// TIA Portal project "EEEB EMBU 4_V17" (V17) (continued)
VERSION : 0.1
   VAR
      "CONNECT-MGE-PCM-E-CF-01" : TCON_IP_v4;   // Dados de configuração
      "CONNECT-MGE-QGBT-AUX-01" : TCON_IP_v4;   // Dados de configuração
      "Register-MGE-PCM-E-CF-01" : Array[0..38] of DInt;   // Tabela para receber os dados
      "Register-MGE-QGBT-AUX-01" : Array[0..38] of DInt;   // Tabela para receber os dados
      LADDR_PROFINET : Hw_IoSystem := 261;   // Endereço de hardware
      MODE_PROFINET : UInt := 4;   // Modo de operação da funcção
      RET_VAL_PROFINET : Int;   // Terorno de diagnóstico
      ESTADO_PROFINET : Array[0..1023] of Bool;   // Diagnóstico da rede PROFINET
      DONE_MB : Array[0..60] of Bool;   // Sinaliza fim de execução
      BUSY_MB : Array[0..60] of Bool;   // Sinaliza espera
      ERROR_MB : Array[0..60] of Bool;   // Sinaliza erro
      STATUS_MB : Array[0..60] of Word;   // Satus da comunicação
      START_MB : Array[0..60] of Bool;   // Inicia comunicação
      FCOM_MB : Array[0..60] of Bool;   // Falha de comunicação
      HAB_MB : Array[0..60] of Bool;   // Habilita comunicação MODBUS
      INICIA_MB : Bool;   // INICIA CICLO DE COMUNICAÇÃO MODBUS
      INI_AUX_MB : Bool;   // AUXILIAR DE INICIALIZAÇÃO
   END_VAR
BEGIN
   "CONNECT-MGE-PCM-E-CF-01".LocalPort := 0;
   "CONNECT-MGE-PCM-E-CF-01".RemotePort := 502;
   "CONNECT-MGE-PCM-E-CF-01".RemoteAddress.ADDR[4] := 59;
   "CONNECT-MGE-PCM-E-CF-01".RemoteAddress.ADDR[3] := 2;
   "CONNECT-MGE-PCM-E-CF-01".RemoteAddress.ADDR[2] := 168;
   "CONNECT-MGE-PCM-E-CF-01".RemoteAddress.ADDR[1] := 192;
   "CONNECT-MGE-PCM-E-CF-01".ActiveEstablished := TRUE;
   "CONNECT-MGE-PCM-E-CF-01".ConnectionType := 11;
   "CONNECT-MGE-PCM-E-CF-01".ID := 10;
   "CONNECT-MGE-PCM-E-CF-01".InterfaceId := 64;
   "CONNECT-MGE-QGBT-AUX-01".LocalPort := 0;
   "CONNECT-MGE-QGBT-AUX-01".RemotePort := 502;
   "CONNECT-MGE-QGBT-AUX-01".RemoteAddress.ADDR[4] := 59;
   "CONNECT-MGE-QGBT-AUX-01".RemoteAddress.ADDR[3] := 2;
   "CONNECT-MGE-QGBT-AUX-01".RemoteAddress.ADDR[2] := 168;
   "CONNECT-MGE-QGBT-AUX-01".RemoteAddress.ADDR[1] := 192;
   "CONNECT-MGE-QGBT-AUX-01".ActiveEstablished := TRUE;
   "CONNECT-MGE-QGBT-AUX-01".ConnectionType := 11;
   "CONNECT-MGE-QGBT-AUX-01".ID := 10;
   "CONNECT-MGE-QGBT-AUX-01".InterfaceId := 64;
   // "Register-MGE-PCM-E-CF-01"[0] : Tensão (L-N) fase 1
   // "Register-MGE-PCM-E-CF-01"[1] : Tensão (L-L) fase 1-2
   // "Register-MGE-PCM-E-CF-01"[2] : Corrente fase 1
   // "Register-MGE-PCM-E-CF-01"[3] : Cos φ fase 1
   // "Register-MGE-PCM-E-CF-01"[4] : Fator de potencia fase 1
   // "Register-MGE-PCM-E-CF-01"[5] : Potencia ativa fase 1
   // "Register-MGE-PCM-E-CF-01"[6] : Potência reativa fase 1
   // "Register-MGE-PCM-E-CF-01"[7] : Potência aparente fase 1
   // "Register-MGE-PCM-E-CF-01"[8] : THDV fase 1
   // "Register-MGE-PCM-E-CF-01"[9] : THDI fase 1
   // "Register-MGE-PCM-E-CF-01"[10] : Tensão (L-N) fase 2
   // "Register-MGE-PCM-E-CF-01"[11] : Tensão (L-L) fase 2-3
   // "Register-MGE-PCM-E-CF-01"[12] : Corrente fase 2
   // "Register-MGE-PCM-E-CF-01"[13] : Cos φ fase 2
   // "Register-MGE-PCM-E-CF-01"[14] : Fator de potência fase 2
   // "Register-MGE-PCM-E-CF-01"[15] : Potência ativa fase 2
   // "Register-MGE-PCM-E-CF-01"[16] : Potência reativa fase 2
   // "Register-MGE-PCM-E-CF-01"[17] : Potência aparente fase 2
   // "Register-MGE-PCM-E-CF-01"[18] : THDV fase 2
   // "Register-MGE-PCM-E-CF-01"[19] : THDI fase 2
   // "Register-MGE-PCM-E-CF-01"[20] : Tensão (L-N) fase 3
   // "Register-MGE-PCM-E-CF-01"[21] : Tensão (L-L) fase 3-1
   // "Register-MGE-PCM-E-CF-01"[22] : Corrente fase 3
   // "Register-MGE-PCM-E-CF-01"[23] : Cos φ fase 3
   // "Register-MGE-PCM-E-CF-01"[24] : Fator de potência fase 3
   // "Register-MGE-PCM-E-CF-01"[25] : Potência ativa fase 3
   // "Register-MGE-PCM-E-CF-01"[26] : Potência reativa fase 3
   // "Register-MGE-PCM-E-CF-01"[27] : Potência aparente fase 3
   // "Register-MGE-PCM-E-CF-01"[28] : THDV fase 3
   // "Register-MGE-PCM-E-CF-01"[29] : THDI fase 3
   // "Register-MGE-PCM-E-CF-01"[30] : Tensão média (L-N)
   // "Register-MGE-PCM-E-CF-01"[31] : Tensão média (L-L)
   // "Register-MGE-PCM-E-CF-01"[32] : Corrente total
   // "Register-MGE-PCM-E-CF-01"[33] : Fator de potência do sistema
   // "Register-MGE-PCM-E-CF-01"[34] : Potência ativa total
   // "Register-MGE-PCM-E-CF-01"[35] : Potência reativa total
   // "Register-MGE-PCM-E-CF-01"[36] : Potência aparente total
   // "Register-MGE-PCM-E-CF-01"[37] : Frequência do sistema
   // "Register-MGE-PCM-E-CF-01"[38] : Corrente de neutro
   // "Register-MGE-QGBT-AUX-01"[37] : Frequência do sistema
   // "Register-MGE-QGBT-AUX-01"[38] : Corrente de neutro
   // "Register-MGE-QGBT-AUX-01"[0] : Tensão (L-N) fase 1
   // "Register-MGE-QGBT-AUX-01"[1] : Tensão (L-L) fase 1-2
   // "Register-MGE-QGBT-AUX-01"[2] : Corrente fase 1
   // "Register-MGE-QGBT-AUX-01"[3] : Cos φ fase 1
   // "Register-MGE-QGBT-AUX-01"[4] : Fator de potencia fase 1
   // "Register-MGE-QGBT-AUX-01"[5] : Potencia ativa fase 1
   // "Register-MGE-QGBT-AUX-01"[6] : Potência reativa fase 1
   // "Register-MGE-QGBT-AUX-01"[7] : Potência aparente fase 1
   // "Register-MGE-QGBT-AUX-01"[8] : THDV fase 1
   // "Register-MGE-QGBT-AUX-01"[9] : THDI fase 1
   // "Register-MGE-QGBT-AUX-01"[10] : Tensão (L-N) fase 2
   // "Register-MGE-QGBT-AUX-01"[11] : Tensão (L-L) fase 2-3
   // "Register-MGE-QGBT-AUX-01"[12] : Corrente fase 2
   // "Register-MGE-QGBT-AUX-01"[13] : Cos φ fase 2
   // "Register-MGE-QGBT-AUX-01"[14] : Fator de potência fase 2
   // "Register-MGE-QGBT-AUX-01"[15] : Potência ativa fase 2
   // "Register-MGE-QGBT-AUX-01"[16] : Potência reativa fase 2
   // "Register-MGE-QGBT-AUX-01"[17] : Potência aparente fase 2
   // "Register-MGE-QGBT-AUX-01"[18] : THDV fase 2
   // "Register-MGE-QGBT-AUX-01"[19] : THDI fase 2
   // "Register-MGE-QGBT-AUX-01"[20] : Tensão (L-N) fase 3
   // "Register-MGE-QGBT-AUX-01"[21] : Tensão (L-L) fase 3-1
   // "Register-MGE-QGBT-AUX-01"[22] : Corrente fase 3
   // "Register-MGE-QGBT-AUX-01"[23] : Cos φ fase 3
   // "Register-MGE-QGBT-AUX-01"[24] : Fator de potência fase 3
   // "Register-MGE-QGBT-AUX-01"[25] : Potência ativa fase 3
   // "Register-MGE-QGBT-AUX-01"[26] : Potência reativa fase 3
   // "Register-MGE-QGBT-AUX-01"[27] : Potência aparente fase 3
   // "Register-MGE-QGBT-AUX-01"[28] : THDV fase 3
   // "Register-MGE-QGBT-AUX-01"[29] : THDI fase 3
   // "Register-MGE-QGBT-AUX-01"[30] : Tensão média (L-N)
   // "Register-MGE-QGBT-AUX-01"[31] : Tensão média (L-L)
   // "Register-MGE-QGBT-AUX-01"[32] : Corrente total
   // "Register-MGE-QGBT-AUX-01"[33] : Fator de potência do sistema
   // "Register-MGE-QGBT-AUX-01"[34] : Potência ativa total
   // "Register-MGE-QGBT-AUX-01"[35] : Potência reativa total
   // "Register-MGE-QGBT-AUX-01"[36] : Potência aparente total
END_DATA_BLOCK

FUNCTION_BLOCK "LOOP"   // FB2, LAD
{ S7_Optimized_Access := 'TRUE' }
VERSION : 0.1
   VAR
      PULSO : Bool;
      AuxLoop : Bool;
      N_L00P : Int;
      Aux_N_LOOP : Int;
      Loop : Int;
   END_VAR
   VAR_TEMP   // added for the SCL form of the ladder/FBD networks
      _w1 : Bool;
      _w2 : Bool;
   END_VAR
BEGIN

REGION Network 2
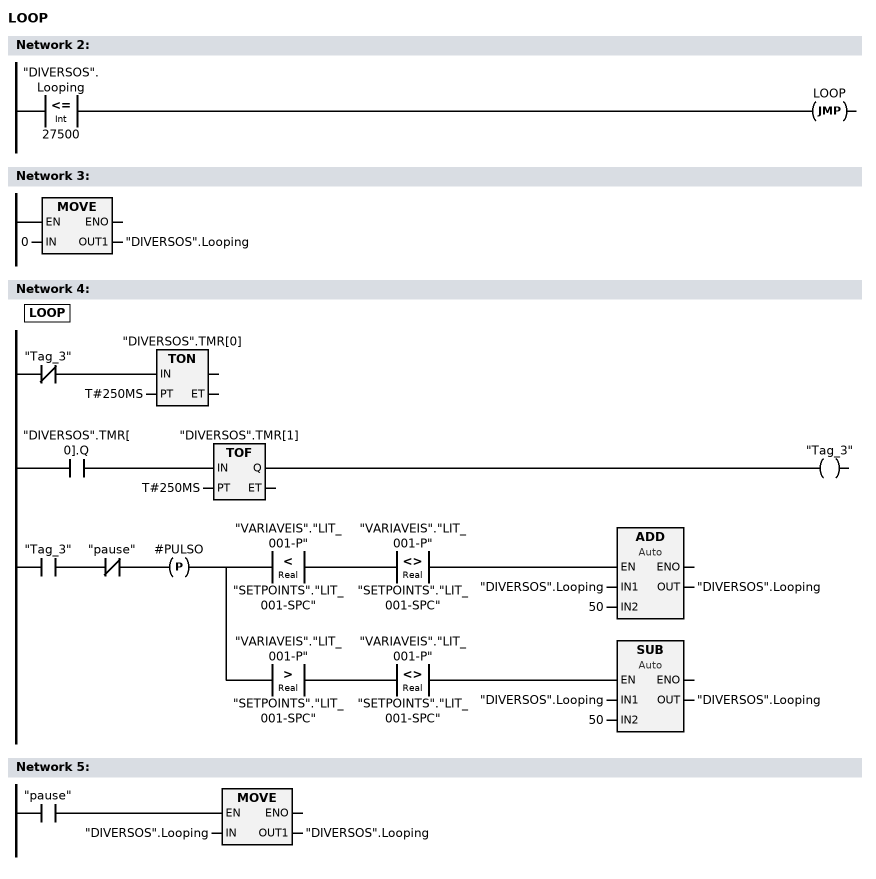
   RUNG wire#powerrail
      { S7_Templates := "SrcType := Int" } LE_Contact(in1 := "DIVERSOS".Looping, in2 := 27500)
      JumpCoil( LOOP )
   END_RUNG
   // the same network as SCL:
   IF "DIVERSOS".Looping <= 27500 THEN GOTO LOOP; END_IF;
END_REGION

REGION Network 3
   RUNG wire#powerrail
      Move(in := 0, out1 => "DIVERSOS".Looping)
   END_RUNG
   // the same network as SCL:
   "DIVERSOS".Looping := 0;
END_REGION

REGION Network 4
   LOOP:
   "DIVERSOS".TMR[0].TON(IN := NOT "Tag_3", PT := T#250MS);
   "DIVERSOS".TMR[1].TOF(IN := "DIVERSOS".TMR[0].Q, PT := T#250MS);
   "Tag_3" := "DIVERSOS".TMR[1].Q;
   #_w1 := "Tag_3" AND NOT "pause";
   #_w2 := #_w1 AND NOT #PULSO;   // rising edge
   #PULSO := #_w1;
   IF #_w2 AND ("VARIAVEIS"."LIT_001-P" < "SETPOINTS"."LIT_001-SPC") AND ("VARIAVEIS"."LIT_001-P" <> "SETPOINTS"."LIT_001-SPC") THEN
       "DIVERSOS".Looping := "DIVERSOS".Looping + 50;
   END_IF;
   IF #_w2 AND ("VARIAVEIS"."LIT_001-P" > "SETPOINTS"."LIT_001-SPC") AND ("VARIAVEIS"."LIT_001-P" <> "SETPOINTS"."LIT_001-SPC") THEN
       "DIVERSOS".Looping := "DIVERSOS".Looping - 50;
   END_IF;
END_REGION

REGION Network 5
   RUNG wire#powerrail
      Contact( "pause" )
      Move(in := "DIVERSOS".Looping, out1 => "DIVERSOS".Looping)
   END_RUNG
   // the same network as SCL:
   IF "pause" THEN "DIVERSOS".Looping := "DIVERSOS".Looping; END_IF;
END_REGION
END_FUNCTION_BLOCK

FUNCTION_BLOCK "ANALOGICOS"   // FB101, LAD
{ S7_Optimized_Access := 'FALSE' }
VERSION : 0.1
   VAR
      LIT_001 : "INSTRUMENTO";   // Nível Tanque
   END_VAR
BEGIN

REGION Network 1: Nível Tanque (Sensor tipo radar)
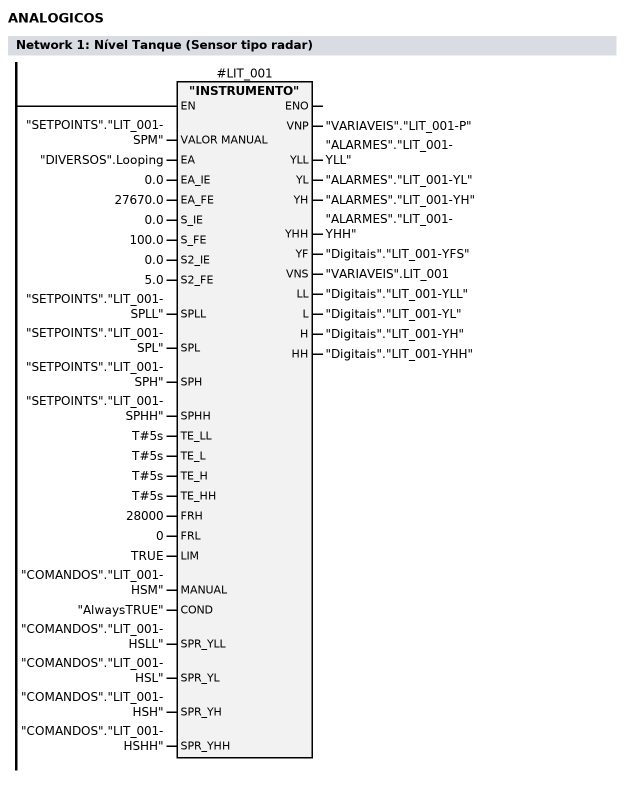
   RUNG wire#powerrail
      #LIT_001("VALOR MANUAL" := "SETPOINTS"."LIT_001-SPM", EA := "DIVERSOS".Looping, EA_IE := 0.0, EA_FE := 27670.0, S_IE := 0.0, S_FE := 100.0, S2_IE := 0.0, S2_FE := 5.0, SPLL := "SETPOINTS"."LIT_001-SPLL", SPL := "SETPOINTS"."LIT_001-SPL", SPH := "SETPOINTS"."LIT_001-SPH", SPHH := "SETPOINTS"."LIT_001-SPHH", TE_LL := T#5s, TE_L := T#5s, TE_H := T#5s, TE_HH := T#5s, FRH := 28000, FRL := 0, LIM := TRUE, MANUAL := "COMANDOS"."LIT_001-HSM", COND := "AlwaysTRUE", SPR_YLL := "COMANDOS"."LIT_001-HSLL", SPR_YL := "COMANDOS"."LIT_001-HSL", SPR_YH := "COMANDOS"."LIT_001-HSH", SPR_YHH := "COMANDOS"."LIT_001-HSHH", VNP => "VARIAVEIS"."LIT_001-P", YLL => "ALARMES"."LIT_001-YLL", YL => "ALARMES"."LIT_001-YL", YH => "ALARMES"."LIT_001-YH", YHH => "ALARMES"."LIT_001-YHH", YF => "Digitais"."LIT_001-YFS", VNS => "VARIAVEIS".LIT_001, LL => "Digitais"."LIT_001-YLL", L => "Digitais"."LIT_001-YL", H => "Digitais"."LIT_001-YH", HH => "Digitais"."LIT_001-YHH")
   END_RUNG
   // the same network as SCL:
   #LIT_001("VALOR MANUAL" := "SETPOINTS"."LIT_001-SPM",   // "INSTRUMENTO"
            EA := "DIVERSOS".Looping,
            EA_IE := 0.0,
            EA_FE := 27670.0,
            S_IE := 0.0,
            S_FE := 100.0,
            S2_IE := 0.0,
            S2_FE := 5.0,
            SPLL := "SETPOINTS"."LIT_001-SPLL",
            SPL := "SETPOINTS"."LIT_001-SPL",
            SPH := "SETPOINTS"."LIT_001-SPH",
            SPHH := "SETPOINTS"."LIT_001-SPHH",
            TE_LL := T#5s,
            TE_L := T#5s,
            TE_H := T#5s,
            TE_HH := T#5s,
            FRH := 28000,
            FRL := 0,
            LIM := TRUE,
            MANUAL := "COMANDOS"."LIT_001-HSM",
            COND := "AlwaysTRUE",
            SPR_YLL := "COMANDOS"."LIT_001-HSLL",
            SPR_YL := "COMANDOS"."LIT_001-HSL",
            SPR_YH := "COMANDOS"."LIT_001-HSH",
            SPR_YHH := "COMANDOS"."LIT_001-HSHH",
            VNP => "VARIAVEIS"."LIT_001-P",
            YLL => "ALARMES"."LIT_001-YLL",
            YL => "ALARMES"."LIT_001-YL",
            YH => "ALARMES"."LIT_001-YH",
            YHH => "ALARMES"."LIT_001-YHH",
            YF => "Digitais"."LIT_001-YFS",
            VNS => "VARIAVEIS".LIT_001,
            LL => "Digitais"."LIT_001-YLL",
            L => "Digitais"."LIT_001-YL",
            H => "Digitais"."LIT_001-YH",
            HH => "Digitais"."LIT_001-YHH");
END_REGION
END_FUNCTION_BLOCK

FUNCTION_BLOCK "MODBUS"   // FB102, LAD
TITLE = BLOCO DE GERENCIAMENTO COMUNICAÇÕES MODBUS/TCP
{ S7_Optimized_Access := 'TRUE' }
VERSION : 0.1
   VAR
      TEFC0 : TON_TIME;   // Tempo para gerar falha de comunicação
      INI_MOD : TON_TIME;   // Tempo para disparar nova comunicação
      TEFC1 : TON_TIME;   // Tempo para gerar falha de comunicação
      TEFC2 : TON_TIME;   // Tempo para gerar falha de comunicação
      TEFC3 : TON_TIME;   // Tempo para gerar falha de comunicação
      TEFC4 : TON_TIME;   // Tempo para gerar falha de comunicação
      TEFC5 : TON_TIME;   // Tempo para gerar falha de comunicação
      TEFC6 : TON_TIME;   // Tempo para gerar falha de comunicação
      TEFC7 : TON_TIME;   // Tempo para gerar falha de comunicação
      TEFC8 : TON_TIME;   // Tempo para gerar falha de comunicação
      TEFC9 : TON_TIME;   // Tempo para gerar falha de comunicação
      TEFC10 : TON_TIME;   // Tempo para gerar falha de comunicação
      TEFC11 : TON_TIME;   // Tempo para gerar falha de comunicação
      TEFC12 : TON_TIME;   // Tempo para gerar falha de comunicação
      TEFC13 : TON_TIME;   // Tempo para gerar falha de comunicação
      TEFC14 : TON_TIME;   // Tempo para gerar falha de comunicação
      TEFC15 : TON_TIME;   // Tempo para gerar falha de comunicação
      TEFC16 : TON_TIME;   // Tempo para gerar falha de comunicação
      TEFC17 : TON_TIME;   // Tempo para gerar falha de comunicação
      TEFC18 : TON_TIME;   // Tempo para gerar falha de comunicação
      TEFC19 : TON_TIME;   // Tempo para gerar falha de comunicação
      TEFC20 : TON_TIME;   // Tempo para gerar falha de comunicação
      TEFC21 : TON_TIME;   // Tempo para gerar falha de comunicação
      TEFC22 : TON_TIME;   // Tempo para gerar falha de comunicação
      TEFC23 : TON_TIME;   // Tempo para gerar falha de comunicação
      TEFC24 : TON_TIME;   // Tempo para gerar falha de comunicação
      TEFC25 : TON_TIME;   // Tempo para gerar falha de comunicação
      TEFC26 : TON_TIME;   // Tempo para gerar falha de comunicação
      TEFC27 : TON_TIME;   // Tempo para gerar falha de comunicação
      TEFC28 : TON_TIME;   // Tempo para gerar falha de comunicação
   END_VAR
BEGIN

REGION Network 1: INICIA LEITURA MODBUS
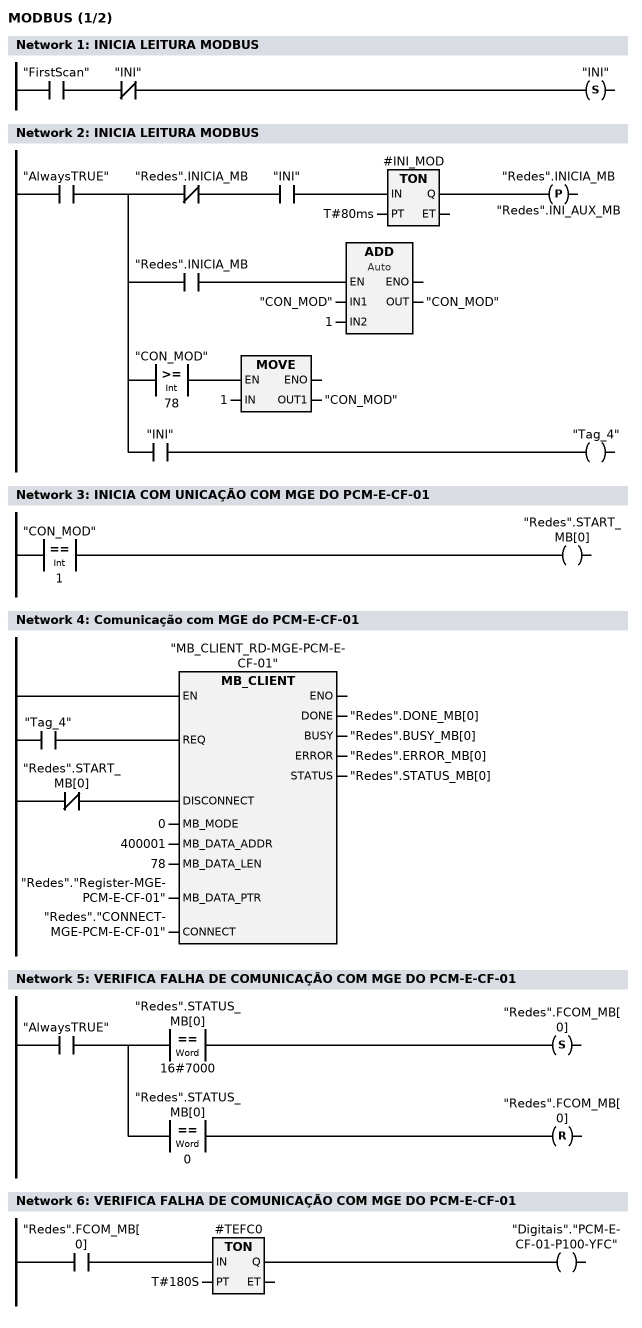
   RUNG wire#powerrail
      Contact( "FirstScan" )
      I_Contact( "INI" )
      S_Coil( "INI" )
   END_RUNG
   // the same network as SCL:
   IF "FirstScan" AND NOT "INI" THEN "INI" := TRUE; END_IF;
END_REGION

REGION Network 2: INICIA LEITURA MODBUS
   #INI_MOD(IN := "AlwaysTRUE" AND NOT "Redes".INICIA_MB AND "INI", PT := T#80ms);   // TON
   "Redes".INICIA_MB := #INI_MOD.Q AND NOT "Redes".INI_AUX_MB;   // rising edge
   "Redes".INI_AUX_MB := #INI_MOD.Q;
   IF "AlwaysTRUE" AND "Redes".INICIA_MB THEN "CON_MOD" := "CON_MOD" + 1; END_IF;
   IF "AlwaysTRUE" AND ("CON_MOD" >= 78) THEN "CON_MOD" := 1; END_IF;
   "Tag_4" := "AlwaysTRUE" AND "INI";
END_REGION

REGION Network 3: INICIA COM UNICAÇÃO COM MGE DO PCM-E-CF-01
   RUNG wire#powerrail
      { S7_Templates := "SrcType := Int" } EQ_Contact(in1 := "CON_MOD", in2 := 1)
      Coil( "Redes".START_MB[0] )
   END_RUNG
   // the same network as SCL:
   "Redes".START_MB[0] := "CON_MOD" = 1;
END_REGION

REGION Network 4: Comunicação com MGE do PCM-E-CF-01
   "MB_CLIENT_RD-MGE-PCM-E-CF-01"(REQ := "Tag_4",   // MB_CLIENT
                           DISCONNECT := NOT "Redes".START_MB[0],
                           MB_MODE := 0,
                           MB_DATA_ADDR := 400001,
                           MB_DATA_LEN := 78,
                           MB_DATA_PTR := "Redes"."Register-MGE-PCM-E-CF-01",
                           CONNECT := "Redes"."CONNECT-MGE-PCM-E-CF-01",
                           DONE => "Redes".DONE_MB[0],
                           BUSY => "Redes".BUSY_MB[0],
                           ERROR => "Redes".ERROR_MB[0],
                           STATUS => "Redes".STATUS_MB[0]);
END_REGION

REGION Network 5: VERIFICA FALHA DE COMUNICAÇÃO COM MGE DO PCM-E-CF-01
   RUNG wire#powerrail
      Contact( "AlwaysTRUE" )
      wire#w1
      { S7_Templates := "SrcType := Word" } EQ_Contact(in1 := "Redes".STATUS_MB[0], in2 := 16#7000)
      S_Coil( "Redes".FCOM_MB[0] )
   END_RUNG
   RUNG wire#w1
      { S7_Templates := "SrcType := Word" } EQ_Contact(in1 := "Redes".STATUS_MB[0], in2 := 0)
      R_Coil( "Redes".FCOM_MB[0] )
   END_RUNG
   // the same network as SCL:
   IF "AlwaysTRUE" AND ("Redes".STATUS_MB[0] = 16#7000) THEN "Redes".FCOM_MB[0] := TRUE; END_IF;
   IF "AlwaysTRUE" AND ("Redes".STATUS_MB[0] = 0) THEN "Redes".FCOM_MB[0] := FALSE; END_IF;
END_REGION

REGION Network 6: VERIFICA FALHA DE COMUNICAÇÃO COM MGE DO PCM-E-CF-01
   #TEFC0(IN := "Redes".FCOM_MB[0], PT := T#180S);   // TON
   "Digitais"."PCM-E-CF-01-P100-YFC" := #TEFC0.Q;
END_REGION

REGION Network 7 (STL): Movimentação de dados do MGE PCM-E-CF-01
   //CONVERSÃO E MOVIMENTAÇÃO MEDIÇÃO DE TENSÃO
         L     "Redes"."Register-MGE-PCM-E-CF-01"[1];
         DTR;
         L     10.0;
         /R;
         T     "VARIAVEIS"."PCM-E-CF-01-04-P100-ETRS";

         L     "Redes"."Register-MGE-PCM-E-CF-01"[11];
         DTR;
         L     10.0;
         /R;
         T     "VARIAVEIS"."PCM-E-CF-01-04-P100-ETST";

         L     "Redes"."Register-MGE-PCM-E-CF-01"[21];
         DTR;
         L     10.0;
         /R;
         T     "VARIAVEIS"."PCM-E-CF-01-04-P100-ETTR";


   //CONVERSÃO E MOVIMENTAÇÃO MEDIÇÃO DE CORRENTE
         L     "Redes"."Register-MGE-PCM-E-CF-01"[2];
         DTR;
         L     100.0;
         /R;
         T     "VARIAVEIS"."PCM-E-CF-01-04-P100-ITR";

         L     "Redes"."Register-MGE-PCM-E-CF-01"[12];
         DTR;
         L     100.0;
         /R;
         T     "VARIAVEIS"."PCM-E-CF-01-04-P100-ITS";

         L     "Redes"."Register-MGE-PCM-E-CF-01"[22];
         DTR;
         L     100.0;
         /R;
         T     "VARIAVEIS"."PCM-E-CF-01-04-P100-ITT";



   //CONVERSÃO E MOVIMENTAÇÃO MEDIÇÃO DE POTÊNCIA ATIVA
         L     "Redes"."Register-MGE-PCM-E-CF-01"[34];
         DTR;
         L     100000.0;
         /R;
         T     "VARIAVEIS"."PCM-E-CF-01-04-P100-JPT";

   //CONVERSÃO E MOVIMENTAÇÃO MEDIÇÃO DE POTÊNCIA REATIVA
         L     "Redes"."Register-MGE-PCM-E-CF-01"[35];
         DTR;
         L     100000.0;
         /R;
         T     "VARIAVEIS"."PCM-E-CF-01-04-P100-JQT";

   //CONVERSÃO E MOVIMENTAÇÃO MEDIÇÃO DE POTÊNCIA APARENTE
         L     "Redes"."Register-MGE-PCM-E-CF-01"[36];
         DTR;
         L     100000.0;
         /R;
         T     "VARIAVEIS"."PCM-E-CF-01-04-P100-JST";

   //CONVERSÃO E MOVIMENTAÇÃO MEDIÇÃO DE FATOR DE POTÊNCIA
         L     %DB500.DBW160;
         ITD;
         DTR;
         L     1000.0;
         /R;
         T     "VARIAVEIS"."PCM-E-CF-01-04-P100-FP";
END_REGION

REGION Network 8: INICIA COM UNICAÇÃO COM MGE DO QGBT-AUX-01
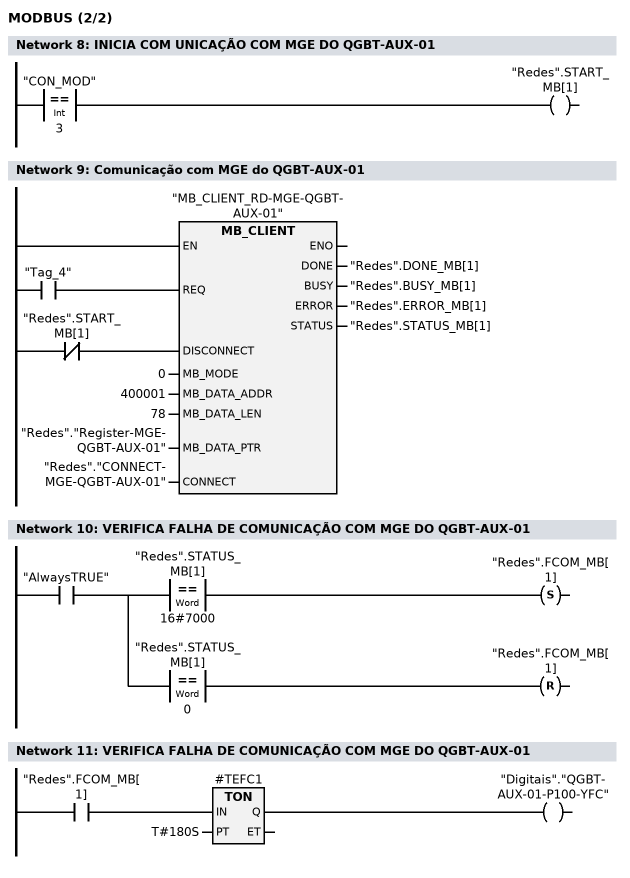
   RUNG wire#powerrail
      { S7_Templates := "SrcType := Int" } EQ_Contact(in1 := "CON_MOD", in2 := 3)
      Coil( "Redes".START_MB[1] )
   END_RUNG
   // the same network as SCL:
   "Redes".START_MB[1] := "CON_MOD" = 3;
END_REGION

REGION Network 9: Comunicação com MGE do QGBT-AUX-01
   "MB_CLIENT_RD-MGE-QGBT-AUX-01"(REQ := "Tag_4",   // MB_CLIENT
                           DISCONNECT := NOT "Redes".START_MB[1],
                           MB_MODE := 0,
                           MB_DATA_ADDR := 400001,
                           MB_DATA_LEN := 78,
                           MB_DATA_PTR := "Redes"."Register-MGE-QGBT-AUX-01",
                           CONNECT := "Redes"."CONNECT-MGE-QGBT-AUX-01",
                           DONE => "Redes".DONE_MB[1],
                           BUSY => "Redes".BUSY_MB[1],
                           ERROR => "Redes".ERROR_MB[1],
                           STATUS => "Redes".STATUS_MB[1]);
END_REGION

REGION Network 10: VERIFICA FALHA DE COMUNICAÇÃO COM MGE DO QGBT-AUX-01
   RUNG wire#powerrail
      Contact( "AlwaysTRUE" )
      wire#w1
      { S7_Templates := "SrcType := Word" } EQ_Contact(in1 := "Redes".STATUS_MB[1], in2 := 16#7000)
      S_Coil( "Redes".FCOM_MB[1] )
   END_RUNG
   RUNG wire#w1
      { S7_Templates := "SrcType := Word" } EQ_Contact(in1 := "Redes".STATUS_MB[1], in2 := 0)
      R_Coil( "Redes".FCOM_MB[1] )
   END_RUNG
   // the same network as SCL:
   IF "AlwaysTRUE" AND ("Redes".STATUS_MB[1] = 16#7000) THEN "Redes".FCOM_MB[1] := TRUE; END_IF;
   IF "AlwaysTRUE" AND ("Redes".STATUS_MB[1] = 0) THEN "Redes".FCOM_MB[1] := FALSE; END_IF;
END_REGION

REGION Network 11: VERIFICA FALHA DE COMUNICAÇÃO COM MGE DO QGBT-AUX-01
   #TEFC1(IN := "Redes".FCOM_MB[1], PT := T#180S);   // TON
   "Digitais"."QGBT-AUX-01-P100-YFC" := #TEFC1.Q;
END_REGION

REGION Network 12 (STL): Movimentação de dados do MGE QGBT-AUX-01
   //CONVERSÃO E MOVIMENTAÇÃO MEDIÇÃO DE TENSÃO
         L     "Redes"."Register-MGE-QGBT-AUX-01"[1];
         DTR;
         L     10.0;
         /R;
         T     "VARIAVEIS"."QGBT-AUX-01-P100-ETRS";

         L     "Redes"."Register-MGE-QGBT-AUX-01"[11];
         DTR;
         L     10.0;
         /R;
         T     "VARIAVEIS"."QGBT-AUX-01-P100-ETST";

         L     "Redes"."Register-MGE-QGBT-AUX-01"[21];
         DTR;
         L     10.0;
         /R;
         T     "VARIAVEIS"."QGBT-AUX-01-P100-ETTR";


   //CONVERSÃO E MOVIMENTAÇÃO MEDIÇÃO DE CORRENTE
         L     "Redes"."Register-MGE-QGBT-AUX-01"[2];
         DTR;
         L     100.0;
         /R;
         T     "VARIAVEIS"."QGBT-AUX-01-P100-ITR";

         L     "Redes"."Register-MGE-QGBT-AUX-01"[12];
         DTR;
         L     100.0;
         /R;
         T     "VARIAVEIS"."QGBT-AUX-01-P100-ITS";

         L     "Redes"."Register-MGE-QGBT-AUX-01"[22];
         DTR;
         L     100.0;
         /R;
         T     "VARIAVEIS"."QGBT-AUX-01-P100-ITT";



   //CONVERSÃO E MOVIMENTAÇÃO MEDIÇÃO DE POTÊNCIA ATIVA
         L     "Redes"."Register-MGE-QGBT-AUX-01"[34];
         DTR;
         L     100000.0;
         /R;
         T     "VARIAVEIS"."QGBT-AUX-01-P100-JPT";

   //CONVERSÃO E MOVIMENTAÇÃO MEDIÇÃO DE POTÊNCIA REATIVA
         L     "Redes"."Register-MGE-QGBT-AUX-01"[35];
         DTR;
         L     100000.0;
         /R;
         T     "VARIAVEIS"."QGBT-AUX-01-P100-JQT";

   //CONVERSÃO E MOVIMENTAÇÃO MEDIÇÃO DE POTÊNCIA APARENTE
         L     "Redes"."Register-MGE-QGBT-AUX-01"[36];
         DTR;
         L     100000.0;
         /R;
         T     "VARIAVEIS"."QGBT-AUX-01-P100-JST";

   //CONVERSÃO E MOVIMENTAÇÃO MEDIÇÃO DE FATOR DE POTÊNCIA
         L     %DB500.DBW316;
         ITD;
         DTR;
         L     1000.0;
         /R;
         T     "VARIAVEIS"."QGBT-AUX-01-P100-FP";
END_REGION
END_FUNCTION_BLOCK

FUNCTION_BLOCK "ROD4"   // FB200, LAD
TITLE = Rodízio de 4 grupos
{ S7_Optimized_Access := 'FALSE' }
VERSION : 0.1
   VAR_INPUT
      G1OK : Bool;   // GRUPO EM CONDIÇÕES DE OPERAÇÃO
      G2OK : Bool;   // GRUPO EM CONDIÇÕES DE OPERAÇÃO
      G3OK : Bool;   // GRUPO EM CONDIÇÕES DE OPERAÇÃO
      G4OK : Bool;   // GRUPO EM CONDIÇÕES DE OPERAÇÃO
      G1L : Bool;   // GRUPO LIGADO
      G2L : Bool;   // GRUPO LIGADO
      G3L : Bool;   // GRUPO LIGADO
      G4L : Bool;   // GRUPO LIGADO
      TEROD : DInt;   // TEMPOPARA RODÍZIO DAS BOMBAS
      LIGP : Bool;   // LIGA BOMBA PRINCIPAL
      LIGC1 : Bool;   // LIGA BOMBA COMPLEMENTAR 1
      LIGC2 : Bool;   // LIGA BOMBA COMPLEMENTAR 2
      LIGC3 : Bool;   // LIGA BOMBA COMPLEMENTAR 3
      DESAB : Bool;   // DESABILITA FUNCIONAMENTO DOS GRUPOS
      T1S : Bool;   // PULSO A CADA 1 SEGUNDO
   END_VAR
   VAR_OUTPUT
      G1P : Bool;   // GRUPO 1 SELECIONADO COMO PRINCIPAL
      G2P : Bool;   // GRUPO 2 SELECIONADO COMO PRINCIPAL
      G3P : Bool;   // GRUPO 3 SELECIONADO COMO PRINCIPAL
      G4P : Bool;   // GRUPO 4 SELECIONADO COMO PRINCIPAL
      G1C1 : Bool;   // GRUPO 1 SELECIONADO COMO COMPLEMENTAR 1
      G2C1 : Bool;   // GRUPO 2 SELECIONADO COMO COMPLEMENTAR 1
      G3C1 : Bool;   // GRUPO 3 SELECIONADO COMO COMPLEMENTAR 1
      G4C1 : Bool;   // GRUPO 4 SELECIONADO COMO COMPLEMENTAR 1
      G1C2 : Bool;   // GRUPO 1 SELECIONADO COMO COMPLEMENTAR 2
      G2C2 : Bool;   // GRUPO 2 SELECIONADO COMO COMPLEMENTAR 2
      G3C2 : Bool;   // GRUPO 3 SELECIONADO COMO COMPLEMENTAR 3
      G4C2 : Bool;   // GRUPO 4 SELECIONADO COMO COMPLEMENTAR 4
      G1C3 : Bool;   // GRUPO 1 SELECIONADO COMO COMPLEMENTAR 3
      G2C3 : Bool;   // GRUPO 2 SELECIONADO COMO COMPLEMENTAR 3
      G3C3 : Bool;   // GRUPO 3 SELECIONADO COMO COMPLEMENTAR 3
      G4C3 : Bool;   // GRUPO 4 SELECIONADO COMO COMPLEMENTAR 3
      LG1 : Bool;   // LIGA GRUPO 1
      LG2 : Bool;   // LIGA GRUPO 2
      LG3 : Bool;   // LIGA GRUPO 3
      LG4 : Bool;   // LIGA GRUPO 4
   END_VAR
   VAR_IN_OUT
      TOG1P : DInt;   // TEMPO DE OPERAÇÃO GRUPO 1
      TOG2P : DInt;   // TEMPO DE OPERAÇÃO GRUPO 2
      TOG3P : DInt;   // TEMPO DE OPERAÇÃO GRUPO 3
      TOG4P : DInt;   // TEMPO DE OPERAÇÃO GRUPO 4
      TEOKG1 : Real;   // TEMPO OK GRUPO 1
      TEOKG2 : Real;   // TEMPO OK GRUPO 2
      TEOKG3 : Real;   // TEMPO OK GRUPO 3
      TEOKG4 : Real;   // TEMPO OK GRUPO 4
   END_VAR
   VAR
      GR1SELP : Bool;   // SELECIONADO COMO PRINCIPAL
      GR2SELP : Bool;   // SELECIONADO COMO PRINCIPAL
      GR3SELP : Bool;   // SELECIONADO COMO PRINCIPAL
      GR4SELP : Bool;   // SELECIONADO COMO PRINCIPAL
      GR1SELC1 : Bool;   // SELECIONADO COMO COMPLEMENTAR 1
      GR2SELC1 : Bool;   // SELECIONADO COMO COMPLEMENTAR 1
      GR3SELC1 : Bool;   // SELECIONADO COMO COMPLEMENTAR 1
      GR4SELC1 : Bool;   // SELECIONADO COMO COMPLEMENTAR 1
      GR1SELC2 : Bool;   // SELECIONADO COMO COMPLEMENTAR 2
      GR2SELC2 : Bool;   // SELECIONADO COMO COMPLEMENTAR 2
      GR3SELC2 : Bool;   // SELECIONADO COMO COMPLEMENTAR 2
      GR4SELC2 : Bool;   // SELECIONADO COMO COMPLEMENTAR 2
      GR1SELC3 : Bool;   // SELECIONADO COMO COMPLEMENTAR 3
      GR2SELC3 : Bool;   // SELECIONADO COMO COMPLEMENTAR 3
      GR3SELC3 : Bool;   // SELECIONADO COMO COMPLEMENTAR 3
      GR4SELC3 : Bool;   // SELECIONADO COMO COMPLEMENTAR 3
      PS1SG1 : Bool;   // AUXILIAR DE PULSO
      PS1SG2 : Bool;   // AUXILIAR DE PULSO
      PS1SG3 : Bool;   // AUXILIAR DE PULSO
      PS1SG4 : Bool;   // AUXILIAR DE PULSO
      PS1 : Bool;   // AUXILIAR DE PULSO
      PS2 : Bool;   // AUXILIAR DE PULSO
      PS3 : Bool;   // AUXILIAR DE PULSO
      PS4 : Bool;   // AUXILIAR DE PULSO
      FIMTEG1 : Bool;   // FIM DO TEMPO DE EXISTÊNCIA DO GRUPO 1
      FIMTEG2 : Bool;   // FIM DO TEMPO DE EXISTÊNCIA DO GRUPO 2
      FIMTEG3 : Bool;   // FIM DO TEMPO DE EXISTÊNCIA DO GRUPO 3
      FIMTEG4 : Bool;   // FIM DO TEMPO DE EXISTÊNCIA DO GRUPO 4
      SDESG1 : Bool;   // SOLICITAÇÃO DE DESLIGAMENTO
      SDESG2 : Bool;   // SOLICITAÇÃO DE DESLIGAMENTO
      SDESG3 : Bool;   // SOLICITAÇÃO DE DESLIGAMENTO
      SDESG4 : Bool;   // SOLICITAÇÃO DE DESLIGAMENTO
      GPL : Bool;   // GRUPO PRINCIPAL LIGADO
      GC1L : Bool;   // GRUPO COMPLEMENTAR 1 LIGADO
      GC2L : Bool;   // GRUPO COMPLEMENTAR 2 LIGADO
      GC3L : Bool;   // GRUPO COMPLEMENTAR 3 LIGADO
      SO_L : Bool;   // SOLICITAÇÃO DE PARTIDA
      SO_D : Bool;   // SOLICITAÇÃO DE DESLIGAMENTO
      RTEOKG1 : Bool;   // RESET TEMPO OK
      RTEOKG2 : Bool;   // RESET TEMPO OK
      RTEOKG3 : Bool;   // RESET TEMPO OK
      RTEOKG4 : Bool;   // RESET TEMPO OK
      TON1 : TON_TIME;   // TEMPORIZADOR
      TON2 : TON_TIME;   // TEMPORIZADOR
      TON3 : TON_TIME;   // TEMPORIZADOR
      TON4 : TON_TIME;   // TEMPORIZADOR
      TSDG1 : TON_TIME;   // TEMPORIZADOR
      TSDG2 : TON_TIME;   // TEMPORIZADOR
      TSDG3 : TON_TIME;   // TEMPORIZADOR
      TSDG4 : TON_TIME;   // TEMPORIZADOR
   END_VAR
   VAR_TEMP
      PRI12 : Bool;   // PRIORIDADE GRUPO 1
      PRI13 : Bool;   // PRIORIDADE GRUPO 1
      PRI14 : Bool;   // PRIORIDADE GRUPO 1
      PRI23 : Bool;   // PRIORIDADE GRUPO 2
      PRI24 : Bool;   // PRIORIDADE GRUPO 2
      PRI34 : Bool;   // PRIORIDADE GRUPO 3
      TMROD : Real;   // TEMPO DE RODIZIO
      NGS : Int;   // NÚMERO DE GRUPOS SOLICITADOS
      NGF : Int;   // NÚMERO DE GRUPOS FUNCIONANDO
      AUX01 : Int;   // AUXILIAR UTILIZADO NA LÓGICA
      AUX02 : Int;   // AUXILIAR UTILIZADO NA LÓGICA
      AUX03 : Int;   // AUXILIAR UTILIZADO NA LÓGICA
      AUX04 : Int;   // AUXILIAR UTILIZADO NA LÓGICA
      AUX05 : Bool;   // AUXILIAR UTILIZADO NA LÓGICA
      AUX06 : Bool;   // AUXILIAR UTILIZADO NA LÓGICA
      AUX07 : Bool;   // AUXILIAR UTILIZADO NA LÓGICA
      AUX08 : Bool;   // AUXILIAR UTILIZADO NA LÓGICA
      ETT1 : Time;   // EFETIVO DO TEMPORIZADOR
      ETT2 : Time;   // EFETIVO DO TEMPORIZADOR
      ETT3 : Time;   // EFETIVO DO TEMPORIZADOR
      ETT4 : Time;   // EFETIVO DO TEMPORIZADOR
      ETTSDG4 : Time;   // EFETIVO DO TEMPORIZADOR
      ETTSDG3 : Time;   // EFETIVO DO TEMPORIZADOR
      ETTSDG2 : Time;   // EFETIVO DO TEMPORIZADOR
      ETTSDG1 : Time;   // EFETIVO DO TEMPORIZADOR
   END_VAR
   VAR_TEMP   // added for the SCL form of the ladder/FBD networks
      _w1 : Bool;
   END_VAR
BEGIN

REGION Network 1: Tranforme em segundo o tempo de rodízio dos sopradores
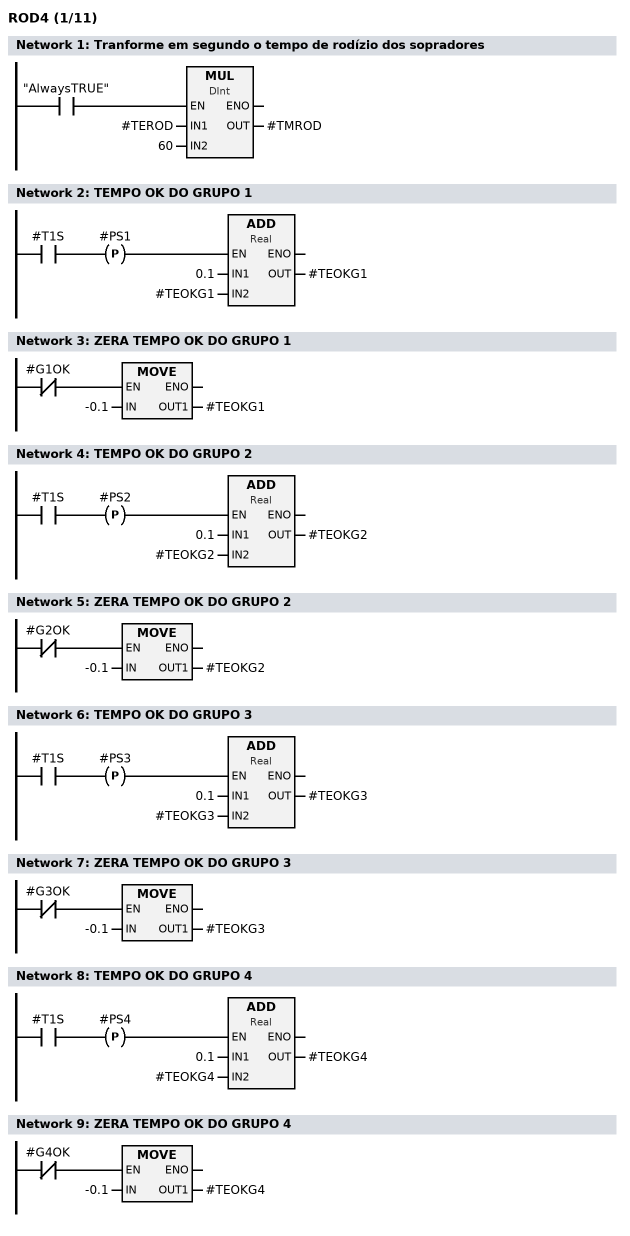
   RUNG wire#powerrail
      Contact( "AlwaysTRUE" )
      { S7_Templates := "SrcType := DInt"; S7_GenerateENO := "TRUE" } Mul(in1 := #TEROD, in2 := 60, out => #TMROD)
   END_RUNG
   // the same network as SCL:
   IF "AlwaysTRUE" THEN #TMROD := #TEROD * 60; END_IF;
END_REGION

REGION Network 2: TEMPO OK DO GRUPO 1
   RUNG wire#powerrail
      Contact( #T1S )
      P_Trig( #PS1 )
      { S7_Templates := "SrcType := Real"; S7_GenerateENO := "TRUE" } Add(in1 := 0.1, in2 := #TEOKG1, out => #TEOKG1)
   END_RUNG
   // the same network as SCL:
   #_w1 := #T1S AND NOT #PS1;   // rising edge
   #PS1 := #T1S;
   IF #_w1 THEN #TEOKG1 := 0.1 + #TEOKG1; END_IF;
END_REGION

REGION Network 3: ZERA TEMPO OK DO GRUPO 1
   RUNG wire#powerrail
      I_Contact( #G1OK )
      { S7_GenerateENO := "TRUE" } Move(in := -0.1, out1 => #TEOKG1)
   END_RUNG
   // the same network as SCL:
   IF NOT #G1OK THEN #TEOKG1 := -0.1; END_IF;
END_REGION

REGION Network 4: TEMPO OK DO GRUPO 2
   RUNG wire#powerrail
      Contact( #T1S )
      P_Trig( #PS2 )
      { S7_Templates := "SrcType := Real"; S7_GenerateENO := "TRUE" } Add(in1 := 0.1, in2 := #TEOKG2, out => #TEOKG2)
   END_RUNG
   // the same network as SCL:
   #_w1 := #T1S AND NOT #PS2;   // rising edge
   #PS2 := #T1S;
   IF #_w1 THEN #TEOKG2 := 0.1 + #TEOKG2; END_IF;
END_REGION

REGION Network 5: ZERA TEMPO OK DO GRUPO 2
   RUNG wire#powerrail
      I_Contact( #G2OK )
      { S7_GenerateENO := "TRUE" } Move(in := -0.1, out1 => #TEOKG2)
   END_RUNG
   // the same network as SCL:
   IF NOT #G2OK THEN #TEOKG2 := -0.1; END_IF;
END_REGION

REGION Network 6: TEMPO OK DO GRUPO 3
   RUNG wire#powerrail
      Contact( #T1S )
      P_Trig( #PS3 )
      { S7_Templates := "SrcType := Real"; S7_GenerateENO := "TRUE" } Add(in1 := 0.1, in2 := #TEOKG3, out => #TEOKG3)
   END_RUNG
   // the same network as SCL:
   #_w1 := #T1S AND NOT #PS3;   // rising edge
   #PS3 := #T1S;
   IF #_w1 THEN #TEOKG3 := 0.1 + #TEOKG3; END_IF;
END_REGION

REGION Network 7: ZERA TEMPO OK DO GRUPO 3
   RUNG wire#powerrail
      I_Contact( #G3OK )
      { S7_GenerateENO := "TRUE" } Move(in := -0.1, out1 => #TEOKG3)
   END_RUNG
   // the same network as SCL:
   IF NOT #G3OK THEN #TEOKG3 := -0.1; END_IF;
END_REGION

REGION Network 8: TEMPO OK DO GRUPO 4
   RUNG wire#powerrail
      Contact( #T1S )
      P_Trig( #PS4 )
      { S7_Templates := "SrcType := Real"; S7_GenerateENO := "TRUE" } Add(in1 := 0.1, in2 := #TEOKG4, out => #TEOKG4)
   END_RUNG
   // the same network as SCL:
   #_w1 := #T1S AND NOT #PS4;   // rising edge
   #PS4 := #T1S;
   IF #_w1 THEN #TEOKG4 := 0.1 + #TEOKG4; END_IF;
END_REGION

REGION Network 9: ZERA TEMPO OK DO GRUPO 4
   RUNG wire#powerrail
      I_Contact( #G4OK )
      { S7_GenerateENO := "TRUE" } Move(in := -0.1, out1 => #TEOKG4)
   END_RUNG
   // the same network as SCL:
   IF NOT #G4OK THEN #TEOKG4 := -0.1; END_IF;
END_REGION

REGION Network 10: DEFINIÇÇÃO DE PRIORIDADE DO GRUPO 1
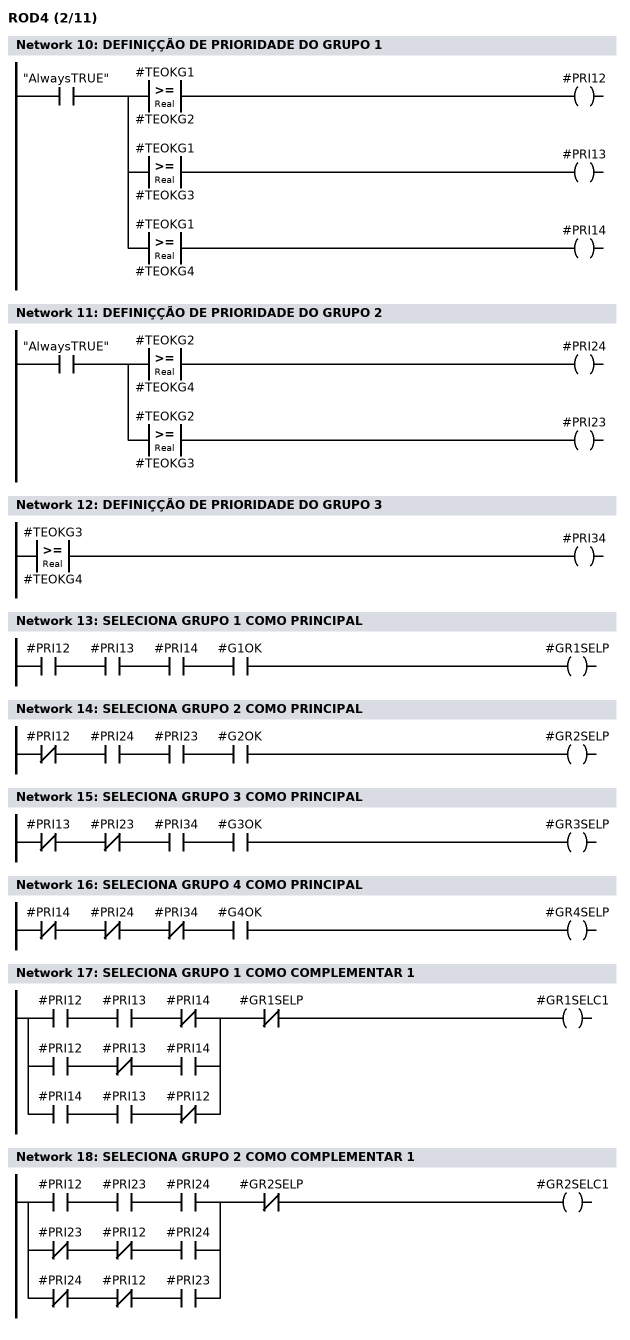
   RUNG wire#powerrail
      Contact( "AlwaysTRUE" )
      wire#w1
      { S7_Templates := "SrcType := Real" } GE_Contact(in1 := #TEOKG1, in2 := #TEOKG2)
      Coil( #PRI12 )
   END_RUNG
   RUNG wire#w1
      { S7_Templates := "SrcType := Real" } GE_Contact(in1 := #TEOKG1, in2 := #TEOKG3)
      Coil( #PRI13 )
   END_RUNG
   RUNG wire#w1
      { S7_Templates := "SrcType := Real" } GE_Contact(in1 := #TEOKG1, in2 := #TEOKG4)
      Coil( #PRI14 )
   END_RUNG
   // the same network as SCL:
   #PRI12 := "AlwaysTRUE" AND (#TEOKG1 >= #TEOKG2);
   #PRI13 := "AlwaysTRUE" AND (#TEOKG1 >= #TEOKG3);
   #PRI14 := "AlwaysTRUE" AND (#TEOKG1 >= #TEOKG4);
END_REGION

REGION Network 11: DEFINIÇÇÃO DE PRIORIDADE DO GRUPO 2
   RUNG wire#powerrail
      Contact( "AlwaysTRUE" )
      wire#w1
      { S7_Templates := "SrcType := Real" } GE_Contact(in1 := #TEOKG2, in2 := #TEOKG4)
      Coil( #PRI24 )
   END_RUNG
   RUNG wire#w1
      { S7_Templates := "SrcType := Real" } GE_Contact(in1 := #TEOKG2, in2 := #TEOKG3)
      Coil( #PRI23 )
   END_RUNG
   // the same network as SCL:
   #PRI24 := "AlwaysTRUE" AND (#TEOKG2 >= #TEOKG4);
   #PRI23 := "AlwaysTRUE" AND (#TEOKG2 >= #TEOKG3);
END_REGION

REGION Network 12: DEFINIÇÇÃO DE PRIORIDADE DO GRUPO 3
   RUNG wire#powerrail
      { S7_Templates := "SrcType := Real" } GE_Contact(in1 := #TEOKG3, in2 := #TEOKG4)
      Coil( #PRI34 )
   END_RUNG
   // the same network as SCL:
   #PRI34 := #TEOKG3 >= #TEOKG4;
END_REGION
